screen "701_Line_Overview_1" 1280x800
   GraphicView "Graphic view_1" at 63,116 size 1157x650; Picture "b1 123927_1"
   Button "Template_Button_3" at 1074,2 size 203x55; TextOn 'FAULT RESET FAULT RESET'; TextOff 'FAULT RESET FAULT RESET'
      on Release: ResetBit("DB_SDC_GLOBAL_M.SDC_ER_Reset")
      on Press: SetBit("DB_SDC_GLOBAL_M.SDC_ER_Reset")
   AlarmView "Template_Alarm view_2" at 128,2 size 948x112
   Button "Template_Button_4" at 1196,56 size 81x59; TextOff 'Text'
      Appearance <- "AlwaysTRUE"
   Button "Button_7" at 0,57 size 128x58; TextOff 'SELECT SCREEN'
      on Release: ActivateScreen("010_START", 0)
   Button "Button_6" at 0,0 size 128x58; TextOff 'PREVIOUS SCREEN'
      on Click: function_efd93a16()
   DateTimeField "Template_Date/time field_2" at 1075,56 size 123x28
   DateTimeField "Template_Date/time field_3" at 1075,83 size 122x32
   TextField "Text field_1" at 981,345 size 46x25; Text 'S14'
   TextField "Text field_2" at 901,345 size 46x25; Text 'S13'
   TextField "Text field_3" at 818,344 size 46x25; Text 'S12'
   TextField "Text field_4" at 778,344 size 46x25; Text 'S11'
   TextField "Text field_5" at 734,344 size 46x25; Text 'S10'
   TextField "Text field_6" at 696,344 size 46x25; Text 'S9'
   TextField "Text field_7" at 653,344 size 46x25; Text 'S57'
   TextField "Text field_8" at 296,344 size 46x25; Text 'S7'
   TextField "Text field_9" at 252,344 size 46x25; Text 'S6'
   TextField "Text field_126" at 454,147 size 327x28; Text 'OVERVIEW 1 - SCREEN 701'
   TextField "Text field_130" at 23,313 size 82x24; Text 'EMS01R2'
   TextField "Text field_131" at 38,329 size 49x24; Text 'JB33'
   TextField "Text field_132" at 28,370 size 71x22; Text 'AREA A'
   TextField "Text field_10" at 135,418 size 46x25; Text 'S5'
   TextField "Text field_11" at 226,507 size 46x25; Text 'S4'
   TextField "Text field_12" at 133,473 size 46x25; Text 'S3'
   TextField "Text field_13" at 13,560 size 46x25; Text 'S2'
   TextField "Text field_14" at 4,640 size 46x25; Text 'S58'
   TextField "Text field_15" at 13,677 size 46x25; Text 'S1'
   TextField "Text field_16" at 5,716 size 46x25; Text 'S56'
   TextField "Text field_17" at 115,721 size 46x25; Text 'S55'
   TextField "Text field_18" at 116,560 size 71x22; Text 'AREA A'
   TextField "Text field_123" at 300,422 size 53x27; Text 'DL1'
   TextField "Text field_116" at 486,494 size 71x22; Text 'AREA G'
   TextField "Text field_119" at 508,426 size 82x22; Text 'AREA AA'
   TextField "Text field_127" at 607,453 size 82x24; Text 'EMS01R3'
   TextField "Text field_129" at 612,518 size 71x22; Text 'AREA B'
   TextField "Text field_19" at 606,485 size 82x22; Text 'AREA AA'
   TextField "Text field_121" at 731,425 size 53x27; Text 'DL2'
   TextField "Text field_122" at 712,450 size 93x25; Text 'Mrg Cell'
   TextField "Text field_120" at 948,425 size 71x22; Text 'AREA B'
   TextField "Text field_20" at 232,731 size 46x25; Text 'S54'
   TextField "Text field_21" at 195,612 size 46x25; Text 'S53'
   TextField "Text field_22" at 278,612 size 46x25; Text 'S52'
   TextField "Text field_23" at 348,613 size 46x25; Text 'S51'
   TextField "Text field_24" at 463,522 size 46x25; Text 'S47'
   TextField "Text field_25" at 534,521 size 46x25; Text 'S48'
   TextField "Text field_26" at 460,696 size 46x25; Text 'S44'
   TextField "Text field_27" at 529,696 size 46x25; Text 'S43'
   TextField "Text field_28" at 667,695 size 46x25; Text 'S42'
   TextField "Text field_29" at 719,657 size 46x25; Text 'S41'
   TextField "Text field_30" at 774,554 size 46x25; Text 'S40'
   TextField "Text field_31" at 883,638 size 46x25; Text 'S39'
   TextField "Text field_32" at 1015,638 size 46x25; Text 'S38'
   TextField "Text field_33" at 1114,638 size 46x25; Text 'S37'
   TextField "Text field_34" at 1158,533 size 46x25; Text 'S36'
   TextField "Text field_35" at 1157,469 size 46x25; Text 'S35'
   TextField "Text field_124" at 109,653 size 49x25; Text 'Cab'
   TextField "Text field_125" at 109,674 size 49x25; Text 'Pick'
   TextField "Text field_117" at 244,698 size 82x22; Text 'AREA FF'
   TextField "Text field_133" at 313,495 size 82x24; Text 'EMS01R1'
   TextField "Text field_134" at 319,518 size 71x22; Text 'AREA G'
   TextField "Text field_135" at 320,545 size 71x22; Text 'AREA F'
   TextField "Text field_136" at 314,570 size 82x22; Text 'AREA FF'
   TextField "Text field_137" at 785,680 size 60x24; Text 'EMS01'
   TextField "Text field_138" at 781,711 size 71x22; Text 'AREA D'
   TextField "Text field_139" at 781,739 size 71x22; Text 'AREA E'
   TextField "Text field_140" at 872,679 size 82x24; Text 'EMS01R4'
   TextField "Text field_143" at 979,672 size 60x24; Text 'EMS01'
   TextField "Text field_144" at 984,686 size 49x24; Text 'JB22'
   TextField "Text field_142" at 878,739 size 71x22; Text 'AREA H'
   TextField "Text field_146" at 973,738 size 71x22; Text 'AREA C'
   TextField "Text field_141" at 872,711 size 82x22; Text 'AREA CC'
   TextField "Text field_145" at 968,710 size 82x22; Text 'AREA BB'
   Button "Button_4" at 3,137 size 127x87; TextOn 'LINE_OVERVIEW_2 LINE OVERVIEW_2'; TextOff 'LINE_OVERVIEW_2 / Main Screen'
      on Click: ActivateScreen("010_START", 0)
   Button "Button_1" at 136,137 size 127x87; TextOn 'LINE_OVERVIEW_2 LINE OVERVIEW_2'; TextOff 'LINE_OVERVIEW_2 System Overview Screen'
      on Click: ActivateScreen("700_System_Line_Overview", 0)
   TextField "Text field_36" at 604,344 size 46x25; Text 'S8'
   Button "Button_2" at 0,0 size 37x32; TextOff 'Text'
      on Release: ActivateScreen("711_CARRIER_STATUS", 0)
      on Press: SetTag("HMI_EMS_Nr", "CarrierNumber")
   Button "Button_5" at 48,712 size 37x32; TextOff 'Text'
      on Release: ActivateScreen("711_CARRIER_STATUS", 0)
      on Press: SetTag("HMI_EMS_Nr", "CarrierNumber")
   Button "Button_8" at 116,760 size 37x32; TextOff 'Text'
      on Release: ActivateScreen("711_CARRIER_STATUS", 0)
      on Press: SetTag("HMI_EMS_Nr", "CarrierNumber")
   Button "Button_9" at 185,729 size 37x32; TextOff 'Text'
      on Release: ActivateScreen("711_CARRIER_STATUS", 0)
      on Press: SetTag("HMI_EMS_Nr", "CarrierNumber")
   Button "Button_10" at 186,691 size 37x32; TextOff 'Text'
      on Release: ActivateScreen("711_CARRIER_STATUS", 0)
      on Press: SetTag("HMI_EMS_Nr", "CarrierNumber")
   Button "Button_11" at 197,654 size 37x32; TextOff 'Text'
      on Release: ActivateScreen("711_CARRIER_STATUS", 0)
      on Press: SetTag("HMI_EMS_Nr", "CarrierNumber")
   Button "Button_12" at 238,654 size 37x32; TextOff 'Text'
      on Release: ActivateScreen("711_CARRIER_STATUS", 0)
      on Press: SetTag("HMI_EMS_Nr", "CarrierNumber")
   Button "Button_13" at 278,654 size 37x32; TextOff 'Text'
      on Release: ActivateScreen("711_CARRIER_STATUS", 0)
      on Press: SetTag("HMI_EMS_Nr", "CarrierNumber")
   Button "Button_14" at 316,654 size 37x32; TextOff 'Text'
      on Release: ActivateScreen("711_CARRIER_STATUS", 0)
      on Press: SetTag("HMI_EMS_Nr", "CarrierNumber")
   Button "Button_15" at 354,654 size 37x32; TextOff 'Text'
      on Release: ActivateScreen("711_CARRIER_STATUS", 0)
      on Press: SetTag("HMI_EMS_Nr", "CarrierNumber")
   Button "Button_16" at 461,654 size 37x32; TextOff 'Text'
      on Release: ActivateScreen("711_CARRIER_STATUS", 0)
      on Press: SetTag("HMI_EMS_Nr", "CarrierNumber")
   Button "Button_17" at 531,654 size 37x32; TextOff 'Text'
      on Release: ActivateScreen("711_CARRIER_STATUS", 0)
      on Press: SetTag("HMI_EMS_Nr", "CarrierNumber")
   Button "Button_18" at 630,654 size 37x32; TextOff 'Text'
      on Release: ActivateScreen("711_CARRIER_STATUS", 0)
      on Press: SetTag("HMI_EMS_Nr", "CarrierNumber")
   Button "Button_19" at 670,654 size 37x32; TextOff 'Text'
      on Release: ActivateScreen("711_CARRIER_STATUS", 0)
      on Press: SetTag("HMI_EMS_Nr", "CarrierNumber")
   Button "Button_20" at 723,623 size 37x32; TextOff 'Text'
      on Release: ActivateScreen("711_CARRIER_STATUS", 0)
      on Press: SetTag("HMI_EMS_Nr", "CarrierNumber")
   Button "Button_21" at 773,599 size 37x32; TextOff 'Text'
      on Release: ActivateScreen("711_CARRIER_STATUS", 0)
      on Press: SetTag("HMI_EMS_Nr", "CarrierNumber")
   Button "Button_22" at 813,599 size 37x32; TextOff 'Text'
      on Release: ActivateScreen("711_CARRIER_STATUS", 0)
      on Press: SetTag("HMI_EMS_Nr", "CarrierNumber")
   Button "Button_23" at 884,599 size 37x32; TextOff 'Text'
      on Release: ActivateScreen("711_CARRIER_STATUS", 0)
      on Press: SetTag("HMI_EMS_Nr", "CarrierNumber")
   Button "Button_24" at 924,599 size 37x32; TextOff 'Text'
      on Release: ActivateScreen("711_CARRIER_STATUS", 0)
      on Press: SetTag("HMI_EMS_Nr", "CarrierNumber")
   Button "Button_25" at 1014,599 size 37x32; TextOff 'Text'
      on Release: ActivateScreen("711_CARRIER_STATUS", 0)
      on Press: SetTag("HMI_EMS_Nr", "CarrierNumber")
   Button "Button_26" at 1054,599 size 37x32; TextOff 'Text'
      on Release: ActivateScreen("711_CARRIER_STATUS", 0)
      on Press: SetTag("HMI_EMS_Nr", "CarrierNumber")
   Button "Button_27" at 1115,599 size 37x32; TextOff 'Text'
      on Release: ActivateScreen("711_CARRIER_STATUS", 0)
      on Press: SetTag("HMI_EMS_Nr", "CarrierNumber")
   Button "Button_28" at 1156,599 size 37x32; TextOff 'Text'
      on Release: ActivateScreen("711_CARRIER_STATUS", 0)
      on Press: SetTag("HMI_EMS_Nr", "CarrierNumber")
   Button "Button_29" at 1218,529 size 37x32; TextOff 'Text'
      on Release: ActivateScreen("711_CARRIER_STATUS", 0)
      on Press: SetTag("HMI_EMS_Nr", "CarrierNumber")
   Button "Button_30" at 1219,466 size 37x32; TextOff 'Text'
      on Release: ActivateScreen("711_CARRIER_STATUS", 0)
      on Press: SetTag("HMI_EMS_Nr", "CarrierNumber")
   Button "Button_31" at 984,371 size 37x32; TextOff 'Text'
      on Release: ActivateScreen("711_CARRIER_STATUS", 0)
      on Press: SetTag("HMI_EMS_Nr", "CarrierNumber")
   Button "Button_32" at 945,371 size 37x32; TextOff 'Text'
      on Release: ActivateScreen("711_CARRIER_STATUS", 0)
      on Press: SetTag("HMI_EMS_Nr", "CarrierNumber")
   Button "Button_33" at 902,371 size 37x32; TextOff 'Text'
      on Release: ActivateScreen("711_CARRIER_STATUS", 0)
      on Press: SetTag("HMI_EMS_Nr", "CarrierNumber")
   Button "Button_34" at 863,371 size 37x32; TextOff 'Text'
      on Release: ActivateScreen("711_CARRIER_STATUS", 0)
      on Press: SetTag("HMI_EMS_Nr", "CarrierNumber")
   Button "Button_35" at 819,371 size 37x32; TextOff 'Text'
      on Release: ActivateScreen("711_CARRIER_STATUS", 0)
      on Press: SetTag("HMI_EMS_Nr", "CarrierNumber")
   Button "Button_36" at 778,371 size 37x32; TextOff 'Text'
      on Release: ActivateScreen("711_CARRIER_STATUS", 0)
      on Press: SetTag("HMI_EMS_Nr", "CarrierNumber")
   Button "Button_37" at 736,371 size 37x32; TextOff 'Text'
      on Release: ActivateScreen("711_CARRIER_STATUS", 0)
      on Press: SetTag("HMI_EMS_Nr", "CarrierNumber")
   Button "Button_38" at 692,371 size 37x32; TextOff 'Text'
      on Release: ActivateScreen("711_CARRIER_STATUS", 0)
      on Press: SetTag("HMI_EMS_Nr", "CarrierNumber")
   Button "Button_39" at 654,371 size 37x32; TextOff 'Text'
      on Release: ActivateScreen("711_CARRIER_STATUS", 0)
      on Press: SetTag("HMI_EMS_Nr", "CarrierNumber")
   Button "Button_40" at 610,371 size 37x32; TextOff 'Text'
      on Release: ActivateScreen("711_CARRIER_STATUS", 0)
      on Press: SetTag("HMI_EMS_Nr", "CarrierNumber")
   Button "Button_41" at 570,371 size 37x32; TextOff 'Text'
      on Release: ActivateScreen("711_CARRIER_STATUS", 0)
      on Press: SetTag("HMI_EMS_Nr", "CarrierNumber")
   Button "Button_42" at 530,371 size 37x32; TextOff 'Text'
      on Release: ActivateScreen("711_CARRIER_STATUS", 0)
      on Press: SetTag("HMI_EMS_Nr", "CarrierNumber")
   Button "Button_43" at 492,371 size 37x32; TextOff 'Text'
      on Release: ActivateScreen("711_CARRIER_STATUS", 0)
      on Press: SetTag("HMI_EMS_Nr", "CarrierNumber")
   Button "Button_44" at 453,371 size 37x32; TextOff 'Text'
      on Release: ActivateScreen("711_CARRIER_STATUS", 0)
      on Press: SetTag("HMI_EMS_Nr", "CarrierNumber")
   Button "Button_45" at 415,371 size 37x32; TextOff 'Text'
      on Release: ActivateScreen("711_CARRIER_STATUS", 0)
      on Press: SetTag("HMI_EMS_Nr", "CarrierNumber")
   Button "Button_46" at 376,371 size 37x32; TextOff 'Text'
      on Release: ActivateScreen("711_CARRIER_STATUS", 0)
      on Press: SetTag("HMI_EMS_Nr", "CarrierNumber")
   Button "Button_47" at 337,371 size 37x32; TextOff 'Text'
      on Release: ActivateScreen("711_CARRIER_STATUS", 0)
      on Press: SetTag("HMI_EMS_Nr", "CarrierNumber")
   Button "Button_48" at 292,371 size 37x32; TextOff 'Text'
      on Release: ActivateScreen("711_CARRIER_STATUS", 0)
      on Press: SetTag("HMI_EMS_Nr", "CarrierNumber")
   Button "Button_49" at 248,371 size 37x32; TextOff 'Text'
      on Release: ActivateScreen("711_CARRIER_STATUS", 0)
      on Press: SetTag("HMI_EMS_Nr", "CarrierNumber")
   Button "Button_50" at 172,414 size 37x32; TextOff 'Text'
      on Release: ActivateScreen("711_CARRIER_STATUS", 0)
      on Press: SetTag("HMI_EMS_Nr", "CarrierNumber")
   Button "Button_51" at 172,449 size 37x32; TextOff 'Text'
      on Release: ActivateScreen("711_CARRIER_STATUS", 0)
      on Press: SetTag("HMI_EMS_Nr", "CarrierNumber")
   Button "Button_52" at 171,503 size 37x32; TextOff 'Text'
      on Release: ActivateScreen("711_CARRIER_STATUS", 0)
      on Press: SetTag("HMI_EMS_Nr", "CarrierNumber")
   Button "Button_53" at 129,503 size 37x32; TextOff 'Text'
      on Release: ActivateScreen("711_CARRIER_STATUS", 0)
      on Press: SetTag("HMI_EMS_Nr", "CarrierNumber")
   TextField "Text field_37" at 579,695 size 46x25; Text 'S63'
   TextField "Text field_38" at 387,613 size 46x25; Text 'S45'
   Button "Button_59" at 584,654 size 37x32; TextOff 'Text'
      on Release: ActivateScreen("711_CARRIER_STATUS", 0)
      on Press: SetTag("HMI_EMS_Nr", "CarrierNumber")
   Group "Group" at 87,503 size 37x32
   Group "Group_1" at 47,596 size 37x32
   Group "Group_2" at 47,635 size 37x32
   Group "Group_3" at 47,672 size 37x32
   Group "Group_4" at 47,555 size 37x32; FormatPattern 99
   Button "Button_60" at 465,556 size 37x32; TextOff 'Text'
      on Release: ActivateScreen("711_CARRIER_STATUS", 0)
      on Press: SetTag("HMI_EMS_Nr", "CarrierNumber")
   Button "Button_61" at 535,556 size 37x32; TextOff 'Text'
      on Release: ActivateScreen("711_CARRIER_STATUS", 0)
      on Press: SetTag("HMI_EMS_Nr", "CarrierNumber")
   Button "Button_58" at 392,654 size 37x32; TextOff 'Text'
      on Release: ActivateScreen("711_CARRIER_STATUS", 0)
      on Press: SetTag("HMI_EMS_Nr", "CarrierNumber")
   IOField "I/O field_30" at 392,654 size 37x32; FormatPattern 99
      ProcessValue <- "CarrierNumber"
      Appearance <- "Faulted"
   IOField "I/O field_8" at 171,503 size 37x32; FormatPattern 99
      ProcessValue <- "CarrierNumber"
      Appearance <- "Faulted"
   IOField "I/O field_11" at 248,371 size 37x32; FormatPattern 99
      ProcessValue <- "CarrierNumber"
      Appearance <- "Faulted"
   IOField "I/O field_12" at 292,371 size 37x32; FormatPattern 99
      ProcessValue <- "CarrierNumber"
      Appearance <- "Faulted"
   IOField "I/O field_13" at 337,371 size 37x32; FormatPattern 99
      ProcessValue <- "CarrierNumber"
      Appearance <- "Faulted"
   IOField "I/O field_14" at 376,371 size 37x32; FormatPattern 99
      ProcessValue <- "CarrierNumber"
      Appearance <- "Faulted"
   IOField "I/O field_15" at 415,371 size 37x32; FormatPattern 99
      ProcessValue <- "CarrierNumber"
      Appearance <- "Faulted"
   IOField "I/O field_16" at 453,371 size 37x32; FormatPattern 99
      ProcessValue <- "CarrierNumber"
      Appearance <- "Faulted"
   IOField "I/O field_17" at 492,371 size 37x32; FormatPattern 99
      ProcessValue <- "CarrierNumber"
      Appearance <- "Faulted"
   IOField "I/O field_18" at 531,371 size 37x32; FormatPattern 99
      ProcessValue <- "CarrierNumber"
      Appearance <- "Faulted"
   IOField "I/O field_19" at 570,371 size 37x32; FormatPattern 99
      ProcessValue <- "CarrierNumber"
      Appearance <- "Faulted"
   IOField "I/O field_20" at 609,371 size 37x32; FormatPattern 99
      ProcessValue <- "CarrierNumber"
      Appearance <- "Faulted"
   IOField "I/O field_21" at 654,371 size 37x32; FormatPattern 99
      ProcessValue <- "CarrierNumber"
   IOField "I/O field_22" at 692,371 size 37x32; FormatPattern 99
      ProcessValue <- "CarrierNumber"
   IOField "I/O field_23" at 736,371 size 37x32; FormatPattern 99
      ProcessValue <- "CarrierNumber"
   IOField "I/O field_24" at 778,371 size 37x32; FormatPattern 99
      ProcessValue <- "CarrierNumber"
   IOField "I/O field_25" at 819,371 size 37x32; FormatPattern 99
      ProcessValue <- "CarrierNumber"
      Appearance <- "Faulted"
   IOField "I/O field_26" at 863,371 size 37x32; FormatPattern 99
      ProcessValue <- "CarrierNumber"
      Appearance <- "Faulted"
   IOField "I/O field_27" at 902,371 size 37x32; FormatPattern 99
      ProcessValue <- "CarrierNumber"
      Appearance <- "Faulted"
   IOField "I/O field_28" at 945,371 size 37x32; FormatPattern 99
      ProcessValue <- "CarrierNumber"
      Appearance <- "Faulted"
   IOField "I/O field_29" at 984,371 size 37x32; FormatPattern 99
      ProcessValue <- "CarrierNumber"
      Appearance <- "Faulted"
   IOField "I/O field_42" at 116,761 size 37x32; FormatPattern 99
      ProcessValue <- "CarrierNumber"
      Appearance <- "Faulted"
   IOField "I/O field_1" at 48,712 size 37x32; FormatPattern 99
      ProcessValue <- "CarrierNumber"
      Appearance <- "Faulted"
   IOField "I/O field_7" at 129,503 size 37x32; FormatPattern 99
      ProcessValue <- "CarrierNumber"
      Appearance <- "Faulted"
   IOField "I/O field_9" at 172,449 size 37x32; FormatPattern 99
      ProcessValue <- "CarrierNumber"
      Appearance <- "Faulted"
   IOField "I/O field_10" at 172,414 size 37x32; FormatPattern 99
      ProcessValue <- "CarrierNumber"
      Appearance <- "Faulted"
   IOField "I/O field_61" at 723,623 size 37x32; FormatPattern 99
      ProcessValue <- "CarrierNumber"
      Appearance <- "Faulted"
   IOField "I/O field_62" at 670,654 size 37x32; FormatPattern 99
      ProcessValue <- "CarrierNumber"
      Appearance <- "Faulted"
   IOField "I/O field_63" at 584,654 size 37x32; FormatPattern 99
      ProcessValue <- "CarrierNumber"
      Appearance <- "Faulted"
   IOField "I/O field_64" at 535,556 size 37x32; FormatPattern 99
      ProcessValue <- "CarrierNumber"
      Appearance <- "Faulted"
   IOField "I/O field_65" at 465,556 size 37x32; FormatPattern 99
      ProcessValue <- "CarrierNumber"
      Appearance <- "Faulted"
   IOField "I/O field_66" at 531,654 size 37x32; FormatPattern 99
      ProcessValue <- "CarrierNumber"
      Appearance <- "Faulted"
   IOField "I/O field_67" at 460,655 size 37x32; FormatPattern 99
      ProcessValue <- "CarrierNumber"
      Appearance <- "Faulted"
   IOField "I/O field_68" at 354,654 size 37x32; FormatPattern 99
      ProcessValue <- "CarrierNumber"
      Appearance <- "Faulted"
   IOField "I/O field_69" at 316,654 size 37x32; FormatPattern 99
      ProcessValue <- "CarrierNumber"
      Appearance <- "Faulted"
   IOField "I/O field_70" at 278,654 size 37x32; FormatPattern 99
      ProcessValue <- "CarrierNumber"
      Appearance <- "Faulted"
   IOField "I/O field_71" at 238,654 size 37x32; FormatPattern 99
      ProcessValue <- "CarrierNumber"
      Appearance <- "Faulted"
   IOField "I/O field_72" at 197,654 size 37x32; FormatPattern 99
      ProcessValue <- "CarrierNumber"
      Appearance <- "Faulted"
   IOField "I/O field_73" at 186,690 size 37x32; FormatPattern 99
      ProcessValue <- "CarrierNumber"
      Appearance <- "Faulted"
   IOField "I/O field_74" at 185,729 size 37x32; FormatPattern 99
      ProcessValue <- "CarrierNumber"
      Appearance <- "Faulted"
   IOField "I/O field_51" at 1219,466 size 37x32; FormatPattern 99
      ProcessValue <- "CarrierNumber"
      Appearance <- "Faulted"
   IOField "I/O field_52" at 1218,529 size 37x32; FormatPattern 99
      ProcessValue <- "CarrierNumber"
      Appearance <- "Faulted"
   IOField "I/O field_53" at 1156,599 size 37x32; FormatPattern 99
      ProcessValue <- "CarrierNumber"
      Appearance <- "Faulted"
   IOField "I/O field_54" at 1115,599 size 37x32; FormatPattern 99
      ProcessValue <- "CarrierNumber"
      Appearance <- "Faulted"
   IOField "I/O field_55" at 1054,599 size 37x32; FormatPattern 99
      ProcessValue <- "CarrierNumber"
      Appearance <- "Faulted"
   IOField "I/O field_56" at 1015,599 size 37x32; FormatPattern 99
      ProcessValue <- "CarrierNumber"
      Appearance <- "Faulted"
   IOField "I/O field_57" at 924,599 size 37x32; FormatPattern 99
      ProcessValue <- "CarrierNumber"
      Appearance <- "Faulted"
   IOField "I/O field_58" at 884,599 size 37x32; FormatPattern 99
      ProcessValue <- "CarrierNumber"
      Appearance <- "Faulted"
   IOField "I/O field_59" at 813,599 size 37x32; FormatPattern 99
      ProcessValue <- "CarrierNumber"
      Appearance <- "Faulted"
   IOField "I/O field_60" at 773,599 size 37x32; FormatPattern 99
      ProcessValue <- "CarrierNumber"
      Appearance <- "Faulted"
   IOField "I/O field_31" at 630,654 size 37x32; FormatPattern 99
      ProcessValue <- "CarrierNumber"
      Appearance <- "Faulted"
   Button "Button_54" at 87,503 size 37x32; TextOff 'Text'
      on Release: ActivateScreen("711_CARRIER_STATUS", 0)
      on Press: SetTag("HMI_EMS_Nr", "CarrierNumber")
   IOField "I/O field_6" at 87,503 size 37x32; FormatPattern 99
      ProcessValue <- "CarrierNumber"
      Appearance <- "Faulted"
   Button "Button_56" at 47,596 size 37x32; TextOff 'Text'
      on Release: ActivateScreen("711_CARRIER_STATUS", 0)
      on Press: SetTag("HMI_EMS_Nr", "CarrierNumber")
   IOField "I/O field_4" at 47,596 size 37x32; FormatPattern 99
      ProcessValue <- "CarrierNumber"
      Appearance <- "Faulted"
   Button "Button_57" at 47,635 size 37x32; TextOff 'Text'
      on Release: ActivateScreen("711_CARRIER_STATUS", 0)
      on Press: SetTag("HMI_EMS_Nr", "CarrierNumber")
   IOField "I/O field_3" at 47,635 size 37x32; FormatPattern 99
      ProcessValue <- "CarrierNumber"
      Appearance <- "Faulted"
   Button "Button_3" at 47,672 size 37x32; TextOff 'Text'
      on Release: ActivateScreen("711_CARRIER_STATUS", 0)
      on Press: SetTag("HMI_EMS_Nr", "CarrierNumber")
   IOField "I/O field_2" at 47,672 size 37x32; FormatPattern 99
      ProcessValue <- "CarrierNumber"
      Appearance <- "Faulted"
   Button "Button_55" at 47,555 size 37x32; TextOff 'Text'
      on Release: ActivateScreen("711_CARRIER_STATUS", 0)
      on Press: SetTag("HMI_EMS_Nr", "CarrierNumber")
   IOField "I/O field_5" at 47,555 size 37x32; FormatPattern 99999
      ProcessValue <- "CarrierNumber"
      Appearance <- "Faulted"

screen "702_Line_Overview_2" 1280x800
   Button "Template_Button_3" at 1074,2 size 203x55; TextOn 'FAULT RESET FAULT RESET'; TextOff 'FAULT RESET FAULT RESET'
      on Release: ResetBit("DB_SDC_GLOBAL_M.SDC_ER_Reset")
      on Press: SetBit("DB_SDC_GLOBAL_M.SDC_ER_Reset")
   AlarmView "Template_Alarm view_2" at 128,2 size 948x112
   Button "Template_Button_4" at 1196,56 size 81x59; TextOff 'Text'
      Appearance <- "AlwaysTRUE"
   Button "Button_7" at 0,57 size 128x58; TextOff 'SELECT SCREEN'
      on Release: ActivateScreen("010_START", 0)
   Button "Button_6" at 0,0 size 128x58; TextOff 'PREVIOUS SCREEN'
      on Click: function_efd93a16()
   DateTimeField "Template_Date/time field_2" at 1075,56 size 123x28
   DateTimeField "Template_Date/time field_3" at 1075,83 size 122x32
   TextField "Text field_2" at 485,123 size 341x28; Text 'OVERVIEW 2 - SCREEN 0024'
   GraphicView "Graphic view_1" at 250,117 size 646x682; Picture "Graphic_3"
   TextField "Text field_1" at 882,117 size 46x25; Text 'S16'
   TextField "Text field_3" at 882,152 size 46x25; Text 'S15'
   TextField "Text field_79" at 605,328 size 60x24; Text 'EMS01'
   TextField "Text field_80" at 608,342 size 49x24; Text 'JB22'
   TextField "Text field_81" at 592,369 size 82x22; Text 'AREA BB'
   TextField "Text field_4" at 477,123 size 327x28; Text 'OVERVIEW 2 - SCREEN 702'
   Button "Button_4" at 1148,702 size 127x87; TextOn 'LINE_OVERVIEW_2 LINE OVERVIEW_2'; TextOff 'LINE_OVERVIEW_2 / Main Screen'
      on Click: ActivateScreen("010_START", 0)
   Button "Button_1" at 1011,702 size 127x87; TextOn 'LINE_OVERVIEW_2 LINE OVERVIEW_2'; TextOff 'LINE_OVERVIEW_2 System Overview Screen'
      on Click: ActivateScreen("700_System_Line_Overview", 0)
   Button "Button_2" at 833,115 size 37x32; TextOff 'Text'
      on Release: ActivateScreen("711_CARRIER_STATUS", 0)
      on Press: SetTag("HMI_EMS_Nr", "CarrierNumber")
   Button "Button_3" at 833,147 size 37x32; TextOff 'Text'
      on Release: ActivateScreen("711_CARRIER_STATUS", 0)
      on Press: SetTag("HMI_EMS_Nr", "CarrierNumber")
   Button "Button_5" at 833,178 size 37x32; TextOff 'Text'
      on Release: ActivateScreen("711_CARRIER_STATUS", 0)
      on Press: SetTag("HMI_EMS_Nr", "CarrierNumber")
   Button "Button_8" at 833,209 size 37x32; TextOff 'Text'
      on Release: ActivateScreen("711_CARRIER_STATUS", 0)
      on Press: SetTag("HMI_EMS_Nr", "CarrierNumber")
   Button "Button_9" at 833,240 size 37x32; TextOff 'Text'
      on Release: ActivateScreen("711_CARRIER_STATUS", 0)
      on Press: SetTag("HMI_EMS_Nr", "CarrierNumber")
   Button "Button_10" at 833,273 size 37x32; TextOff 'Text'
      on Release: ActivateScreen("711_CARRIER_STATUS", 0)
      on Press: SetTag("HMI_EMS_Nr", "CarrierNumber")
   Button "Button_11" at 833,305 size 37x32; TextOff 'Text'
      on Release: ActivateScreen("711_CARRIER_STATUS", 0)
      on Press: SetTag("HMI_EMS_Nr", "CarrierNumber")
   Button "Button_12" at 833,337 size 37x32; TextOff 'Text'
      on Release: ActivateScreen("711_CARRIER_STATUS", 0)
      on Press: SetTag("HMI_EMS_Nr", "CarrierNumber")
   Button "Button_13" at 833,369 size 37x32; TextOff 'Text'
      on Release: ActivateScreen("711_CARRIER_STATUS", 0)
      on Press: SetTag("HMI_EMS_Nr", "CarrierNumber")
   Button "Button_14" at 833,401 size 37x32; TextOff 'Text'
      on Release: ActivateScreen("711_CARRIER_STATUS", 0)
      on Press: SetTag("HMI_EMS_Nr", "CarrierNumber")
   Button "Button_15" at 833,433 size 37x32; TextOff 'Text'
      on Release: ActivateScreen("711_CARRIER_STATUS", 0)
      on Press: SetTag("HMI_EMS_Nr", "CarrierNumber")
   Button "Button_16" at 833,464 size 37x32; TextOff 'Text'
      on Release: ActivateScreen("711_CARRIER_STATUS", 0)
      on Press: SetTag("HMI_EMS_Nr", "CarrierNumber")
   Button "Button_17" at 833,496 size 37x32; TextOff 'Text'
      on Release: ActivateScreen("711_CARRIER_STATUS", 0)
      on Press: SetTag("HMI_EMS_Nr", "CarrierNumber")
   Button "Button_18" at 833,528 size 37x32; TextOff 'Text'
      on Release: ActivateScreen("711_CARRIER_STATUS", 0)
      on Press: SetTag("HMI_EMS_Nr", "CarrierNumber")
   Button "Button_19" at 833,560 size 37x32; TextOff 'Text'
      on Release: ActivateScreen("711_CARRIER_STATUS", 0)
      on Press: SetTag("HMI_EMS_Nr", "CarrierNumber")
   Button "Button_20" at 833,592 size 37x32; TextOff 'Text'
      on Release: ActivateScreen("711_CARRIER_STATUS", 0)
      on Press: SetTag("HMI_EMS_Nr", "CarrierNumber")
   Button "Button_21" at 833,623 size 37x32; TextOff 'Text'
      on Release: ActivateScreen("711_CARRIER_STATUS", 0)
      on Press: SetTag("HMI_EMS_Nr", "CarrierNumber")
   Button "Button_22" at 833,654 size 37x32; TextOff 'Text'
      on Release: ActivateScreen("711_CARRIER_STATUS", 0)
      on Press: SetTag("HMI_EMS_Nr", "CarrierNumber")
   Button "Button_23" at 833,686 size 37x32; TextOff 'Text'
      on Release: ActivateScreen("711_CARRIER_STATUS", 0)
      on Press: SetTag("HMI_EMS_Nr", "CarrierNumber")
   Button "Button_24" at 833,718 size 37x32; TextOff 'Text'
      on Release: ActivateScreen("711_CARRIER_STATUS", 0)
      on Press: SetTag("HMI_EMS_Nr", "CarrierNumber")
   Button "Button_25" at 833,750 size 37x32; TextOff 'Text'
      on Release: ActivateScreen("711_CARRIER_STATUS", 0)
      on Press: SetTag("HMI_EMS_Nr", "CarrierNumber")
   IOField "I/O field_30" at 833,750 size 37x32; FormatPattern 99
      ProcessValue <- "CarrierNumber"
      Appearance <- "Faulted"
   IOField "I/O field_31" at 833,718 size 37x32; FormatPattern 99
      ProcessValue <- "CarrierNumber"
      Appearance <- "Faulted"
   IOField "I/O field_32" at 833,686 size 37x32; FormatPattern 99
      ProcessValue <- "CarrierNumber"
      Appearance <- "Faulted"
   IOField "I/O field_33" at 833,654 size 37x32; FormatPattern 99
      ProcessValue <- "CarrierNumber"
      Appearance <- "Faulted"
   IOField "I/O field_34" at 833,623 size 37x32; FormatPattern 99
      ProcessValue <- "CarrierNumber"
      Appearance <- "Faulted"
   IOField "I/O field_35" at 833,592 size 37x32; FormatPattern 99
      ProcessValue <- "CarrierNumber"
      Appearance <- "Faulted"
   IOField "I/O field_36" at 833,560 size 37x32; FormatPattern 99
      ProcessValue <- "CarrierNumber"
      Appearance <- "Faulted"
   IOField "I/O field_37" at 833,528 size 37x32; FormatPattern 99
      ProcessValue <- "CarrierNumber"
      Appearance <- "Faulted"
   IOField "I/O field_38" at 833,496 size 37x32; FormatPattern 99
      ProcessValue <- "CarrierNumber"
      Appearance <- "Faulted"
   IOField "I/O field_39" at 833,464 size 37x32; FormatPattern 99
      ProcessValue <- "CarrierNumber"
      Appearance <- "Faulted"
   IOField "I/O field_55" at 833,114 size 37x32; FormatPattern 99
      ProcessValue <- "CarrierNumber"
      Appearance <- "Faulted"
   IOField "I/O field_56" at 833,146 size 37x32; FormatPattern 99
      ProcessValue <- "CarrierNumber"
      Appearance <- "Faulted"
   IOField "I/O field_57" at 833,177 size 37x32; FormatPattern 99
      ProcessValue <- "CarrierNumber"
      Appearance <- "Faulted"
   IOField "I/O field_58" at 833,209 size 37x32; FormatPattern 99
      ProcessValue <- "CarrierNumber"
      Appearance <- "Faulted"
   IOField "I/O field_59" at 833,241 size 37x32; FormatPattern 99
      ProcessValue <- "CarrierNumber"
      Appearance <- "Faulted"
   IOField "I/O field_60" at 833,273 size 37x32; FormatPattern 99
      ProcessValue <- "CarrierNumber"
      Appearance <- "Faulted"
   IOField "I/O field_61" at 833,305 size 37x32; FormatPattern 99
      ProcessValue <- "CarrierNumber"
      Appearance <- "Faulted"
   IOField "I/O field_62" at 833,337 size 37x32; FormatPattern 99
      ProcessValue <- "CarrierNumber"
      Appearance <- "Faulted"
   IOField "I/O field_63" at 833,369 size 37x32; FormatPattern 99
      ProcessValue <- "CarrierNumber"
      Appearance <- "Faulted"
   IOField "I/O field_64" at 833,401 size 37x32; FormatPattern 99
      ProcessValue <- "CarrierNumber"
      Appearance <- "Faulted"
   IOField "I/O field_65" at 833,433 size 37x32; FormatPattern 99
      ProcessValue <- "CarrierNumber"
      Appearance <- "Faulted"

screen "703_Line_Overview_3" 1280x800
   Button "Template_Button_3" at 1074,2 size 203x55; TextOn 'FAULT RESET FAULT RESET'; TextOff 'FAULT RESET FAULT RESET'
      on Release: ResetBit("DB_SDC_GLOBAL_M.SDC_ER_Reset")
      on Press: SetBit("DB_SDC_GLOBAL_M.SDC_ER_Reset")
   AlarmView "Template_Alarm view_2" at 128,2 size 948x112
   Button "Template_Button_4" at 1196,56 size 81x59; TextOff 'Text'
      Appearance <- "AlwaysTRUE"
   Button "Button_7" at 0,57 size 128x58; TextOff 'SELECT SCREEN'
      on Release: ActivateScreen("010_START", 0)
   Button "Button_6" at 0,0 size 128x58; TextOff 'PREVIOUS SCREEN'
      on Click: function_efd93a16()
   DateTimeField "Template_Date/time field_2" at 1075,56 size 123x28
   DateTimeField "Template_Date/time field_3" at 1075,83 size 122x32
   GraphicView "Graphic view_1" at 26,247 size 1142x552; Picture "b2 124337_2"
   TextField "Text field_1" at 910,378 size 46x25; Text 'S17'
   TextField "Text field_15" at 77,290 size 46x25; Text 'S21'
   TextField "Text field_16" at 209,383 size 46x25; Text 'S20'
   TextField "Text field_17" at 612,381 size 46x25; Text 'S19'
   TextField "Text field_18" at 752,380 size 46x25; Text 'S18'
   TextField "Text field_5" at 1038,197 size 46x25; Text 'S32'
   TextField "Text field_6" at 828,197 size 46x25; Text 'S31'
   TextField "Text field_7" at 663,197 size 46x25; Text 'S30'
   TextField "Text field_8" at 577,197 size 46x25; Text 'S29'
   TextField "Text field_9" at 491,197 size 46x25; Text 'S28'
   TextField "Text field_10" at 414,197 size 46x25; Text 'S27'
   TextField "Text field_11" at 339,197 size 46x25; Text 'S26'
   TextField "Text field_12" at 277,163 size 46x25; Text 'S24'
   TextField "Text field_13" at 276,276 size 46x25; Text 'S23'
   TextField "Text field_14" at 211,198 size 46x25; Text 'S22'
   TextField "Text field_2" at 485,123 size 327x28; Text 'OVERVIEW 3 - SCREEN 703'
   TextField "Text field_4" at 1116,767 size 46x25; Text 'S33'
   TextField "Text field_79" at 1009,409 size 60x24; Text 'EMS01'
   TextField "Text field_80" at 1012,423 size 49x24; Text 'JB22'
   TextField "Text field_82" at 1002,461 size 71x22; Text 'AREA C'
   TextField "Text field_3" at 738,426 size 71x22; Text 'AREA C'
   TextField "Text field_76" at 379,430 size 82x24; Text 'EMS01R4'
   TextField "Text field_77" at 378,459 size 82x22; Text 'AREA CC'
   TextField "Text field_78" at 383,487 size 71x22; Text 'AREA H'
   TextField "Text field_73" at 123,291 size 82x22; Text 'AREA CC'
   TextField "Text field_121" at 489,285 size 61x28; Text 'DL5'
   TextField "Text field_72" at 926,291 size 71x22; Text 'AREA H'
   TextField "Text field_71" at 1077,550 size 71x22; Text 'AREA D'
   TextField "Text field_93" at 1008,626 size 60x24; Text 'EMS01'
   TextField "Text field_94" at 1003,660 size 71x22; Text 'AREA D'
   Button "Button_4" at 26,689 size 127x87; TextOn 'LINE_OVERVIEW_2 LINE OVERVIEW_2'; TextOff 'LINE_OVERVIEW_2 / Main Screen'
      on Click: ActivateScreen("010_START", 0)
   Button "Button_1" at 158,689 size 127x87; TextOn 'LINE_OVERVIEW_2 LINE OVERVIEW_2'; TextOff 'LINE_OVERVIEW_2 System Overview Screen'
      on Click: ActivateScreen("700_System_Line_Overview", 0)
   Button "Button_2" at 855,532 size 37x32; TextOff 'Text'
      on Release: ActivateScreen("711_CARRIER_STATUS", 0)
      on Press: SetTag("HMI_EMS_Nr", "CarrierNumber")
   Button "Button_3" at 855,500 size 37x32; TextOff 'Text'
      on Release: ActivateScreen("711_CARRIER_STATUS", 0)
      on Press: SetTag("HMI_EMS_Nr", "CarrierNumber")
   Button "Button_5" at 855,467 size 37x32; TextOff 'Text'
      on Release: ActivateScreen("711_CARRIER_STATUS", 0)
      on Press: SetTag("HMI_EMS_Nr", "CarrierNumber")
   Button "Button_8" at 855,435 size 37x32; TextOff 'Text'
      on Release: ActivateScreen("711_CARRIER_STATUS", 0)
      on Press: SetTag("HMI_EMS_Nr", "CarrierNumber")
   Button "Button_9" at 855,404 size 37x32; TextOff 'Text'
      on Release: ActivateScreen("711_CARRIER_STATUS", 0)
      on Press: SetTag("HMI_EMS_Nr", "CarrierNumber")
   Button "Button_10" at 855,372 size 37x32; TextOff 'Text'
      on Release: ActivateScreen("711_CARRIER_STATUS", 0)
      on Press: SetTag("HMI_EMS_Nr", "CarrierNumber")
   Button "Button_11" at 799,343 size 37x32; TextOff 'Text'
      on Release: ActivateScreen("711_CARRIER_STATUS", 0)
      on Press: SetTag("HMI_EMS_Nr", "CarrierNumber")
   Button "Button_12" at 753,343 size 37x32; TextOff 'Text'
      on Release: ActivateScreen("711_CARRIER_STATUS", 0)
      on Press: SetTag("HMI_EMS_Nr", "CarrierNumber")
   Button "Button_13" at 661,344 size 37x32; TextOff 'Text'
      on Release: ActivateScreen("711_CARRIER_STATUS", 0)
      on Press: SetTag("HMI_EMS_Nr", "CarrierNumber")
   Button "Button_14" at 613,344 size 37x32; TextOff 'Text'
      on Release: ActivateScreen("711_CARRIER_STATUS", 0)
      on Press: SetTag("HMI_EMS_Nr", "CarrierNumber")
   Button "Button_15" at 519,344 size 37x32; TextOff 'Text'
      on Release: ActivateScreen("711_CARRIER_STATUS", 0)
      on Press: SetTag("HMI_EMS_Nr", "CarrierNumber")
   Button "Button_16" at 475,344 size 37x32; TextOff 'Text'
      on Release: ActivateScreen("711_CARRIER_STATUS", 0)
      on Press: SetTag("HMI_EMS_Nr", "CarrierNumber")
   Button "Button_17" at 431,344 size 37x32; TextOff 'Text'
      on Release: ActivateScreen("711_CARRIER_STATUS", 0)
      on Press: SetTag("HMI_EMS_Nr", "CarrierNumber")
   Button "Button_18" at 387,344 size 37x32; TextOff 'Text'
      on Release: ActivateScreen("711_CARRIER_STATUS", 0)
      on Press: SetTag("HMI_EMS_Nr", "CarrierNumber")
   Button "Button_19" at 343,344 size 37x32; TextOff 'Text'
      on Release: ActivateScreen("711_CARRIER_STATUS", 0)
      on Press: SetTag("HMI_EMS_Nr", "CarrierNumber")
   Button "Button_20" at 299,344 size 37x32; TextOff 'Text'
      on Release: ActivateScreen("711_CARRIER_STATUS", 0)
      on Press: SetTag("HMI_EMS_Nr", "CarrierNumber")
   Button "Button_21" at 255,344 size 37x32; TextOff 'Text'
      on Release: ActivateScreen("711_CARRIER_STATUS", 0)
      on Press: SetTag("HMI_EMS_Nr", "CarrierNumber")
   Button "Button_22" at 211,344 size 37x32; TextOff 'Text'
      on Release: ActivateScreen("711_CARRIER_STATUS", 0)
      on Press: SetTag("HMI_EMS_Nr", "CarrierNumber")
   Button "Button_23" at 17,285 size 37x32; TextOff 'Text'
      on Release: ActivateScreen("711_CARRIER_STATUS", 0)
      on Press: SetTag("HMI_EMS_Nr", "CarrierNumber")
   Button "Button_24" at 122,230 size 37x32; TextOff 'Text'
      on Release: ActivateScreen("711_CARRIER_STATUS", 0)
      on Press: SetTag("HMI_EMS_Nr", "CarrierNumber")
   Button "Button_25" at 166,230 size 37x32; TextOff 'Text'
      on Release: ActivateScreen("711_CARRIER_STATUS", 0)
      on Press: SetTag("HMI_EMS_Nr", "CarrierNumber")
   Button "Button_26" at 212,230 size 37x32; TextOff 'Text'
      on Release: ActivateScreen("711_CARRIER_STATUS", 0)
      on Press: SetTag("HMI_EMS_Nr", "CarrierNumber")
   Button "Button_27" at 278,230 size 37x32; TextOff 'Text'
      on Release: ActivateScreen("711_CARRIER_STATUS", 0)
      on Press: SetTag("HMI_EMS_Nr", "CarrierNumber")
   Button "Button_28" at 342,230 size 37x32; TextOff 'Text'
      on Release: ActivateScreen("711_CARRIER_STATUS", 0)
      on Press: SetTag("HMI_EMS_Nr", "CarrierNumber")
   Button "Button_29" at 415,230 size 37x32; TextOff 'Text'
      on Release: ActivateScreen("711_CARRIER_STATUS", 0)
      on Press: SetTag("HMI_EMS_Nr", "CarrierNumber")
   Button "Button_30" at 279,193 size 37x32; TextOff 'Text'
      on Release: ActivateScreen("711_CARRIER_STATUS", 0)
      on Press: SetTag("HMI_EMS_Nr", "CarrierNumber")
   Button "Button_31" at 492,230 size 37x32; TextOff 'Text'
      on Release: ActivateScreen("711_CARRIER_STATUS", 0)
      on Press: SetTag("HMI_EMS_Nr", "CarrierNumber")
   Button "Button_32" at 578,230 size 37x32; TextOff 'Text'
      on Release: ActivateScreen("711_CARRIER_STATUS", 0)
      on Press: SetTag("HMI_EMS_Nr", "CarrierNumber")
   Button "Button_33" at 665,230 size 37x32; TextOff 'Text'
      on Release: ActivateScreen("711_CARRIER_STATUS", 0)
      on Press: SetTag("HMI_EMS_Nr", "CarrierNumber")
   Button "Button_34" at 768,230 size 37x32; TextOff 'Text'
      on Release: ActivateScreen("711_CARRIER_STATUS", 0)
      on Press: SetTag("HMI_EMS_Nr", "CarrierNumber")
   Button "Button_35" at 831,230 size 37x32; TextOff 'Text'
      on Release: ActivateScreen("711_CARRIER_STATUS", 0)
      on Press: SetTag("HMI_EMS_Nr", "CarrierNumber")
   Button "Button_36" at 974,230 size 37x32; TextOff 'Text'
      on Release: ActivateScreen("711_CARRIER_STATUS", 0)
      on Press: SetTag("HMI_EMS_Nr", "CarrierNumber")
   Button "Button_37" at 1041,230 size 37x32; TextOff 'Text'
      on Release: ActivateScreen("711_CARRIER_STATUS", 0)
      on Press: SetTag("HMI_EMS_Nr", "CarrierNumber")
   Button "Button_38" at 1174,267 size 37x32; TextOff 'Text'
      on Release: ActivateScreen("711_CARRIER_STATUS", 0)
      on Press: SetTag("HMI_EMS_Nr", "CarrierNumber")
   Button "Button_39" at 1174,300 size 37x32; TextOff 'Text'
      on Release: ActivateScreen("711_CARRIER_STATUS", 0)
      on Press: SetTag("HMI_EMS_Nr", "CarrierNumber")
   Button "Button_40" at 1174,333 size 37x32; TextOff 'Text'
      on Release: ActivateScreen("711_CARRIER_STATUS", 0)
      on Press: SetTag("HMI_EMS_Nr", "CarrierNumber")
   Button "Button_41" at 1174,366 size 37x32; TextOff 'Text'
      on Release: ActivateScreen("711_CARRIER_STATUS", 0)
      on Press: SetTag("HMI_EMS_Nr", "CarrierNumber")
   Button "Button_42" at 1174,399 size 37x32; TextOff 'Text'
      on Release: ActivateScreen("711_CARRIER_STATUS", 0)
      on Press: SetTag("HMI_EMS_Nr", "CarrierNumber")
   Button "Button_43" at 1174,432 size 37x32; TextOff 'Text'
      on Release: ActivateScreen("711_CARRIER_STATUS", 0)
      on Press: SetTag("HMI_EMS_Nr", "CarrierNumber")
   Button "Button_44" at 1174,465 size 37x32; TextOff 'Text'
      on Release: ActivateScreen("711_CARRIER_STATUS", 0)
      on Press: SetTag("HMI_EMS_Nr", "CarrierNumber")
   Button "Button_45" at 1174,498 size 37x32; TextOff 'Text'
      on Release: ActivateScreen("711_CARRIER_STATUS", 0)
      on Press: SetTag("HMI_EMS_Nr", "CarrierNumber")
   Button "Button_46" at 1174,531 size 37x32; TextOff 'Text'
      on Release: ActivateScreen("711_CARRIER_STATUS", 0)
      on Press: SetTag("HMI_EMS_Nr", "CarrierNumber")
   Button "Button_47" at 1174,564 size 37x32; TextOff 'Text'
      on Release: ActivateScreen("711_CARRIER_STATUS", 0)
      on Press: SetTag("HMI_EMS_Nr", "CarrierNumber")
   Button "Button_48" at 1174,597 size 37x32; TextOff 'Text'
      on Release: ActivateScreen("711_CARRIER_STATUS", 0)
      on Press: SetTag("HMI_EMS_Nr", "CarrierNumber")
   Button "Button_49" at 1174,630 size 37x32; TextOff 'Text'
      on Release: ActivateScreen("711_CARRIER_STATUS", 0)
      on Press: SetTag("HMI_EMS_Nr", "CarrierNumber")
   Button "Button_50" at 1174,663 size 37x32; TextOff 'Text'
      on Release: ActivateScreen("711_CARRIER_STATUS", 0)
      on Press: SetTag("HMI_EMS_Nr", "CarrierNumber")
   Button "Button_51" at 1174,696 size 37x32; TextOff 'Text'
      on Release: ActivateScreen("711_CARRIER_STATUS", 0)
      on Press: SetTag("HMI_EMS_Nr", "CarrierNumber")
   Button "Button_52" at 1174,729 size 37x32; TextOff 'Text'
      on Release: ActivateScreen("711_CARRIER_STATUS", 0)
      on Press: SetTag("HMI_EMS_Nr", "CarrierNumber")
   Button "Button_53" at 1174,762 size 37x32; TextOff 'Text'
      on Release: ActivateScreen("711_CARRIER_STATUS", 0)
      on Press: SetTag("HMI_EMS_Nr", "CarrierNumber")
   IOField "I/O field_3" at 17,285 size 37x32; FormatPattern 99
      ProcessValue <- "CarrierNumber"
      Appearance <- "Faulted"
   IOField "I/O field_37" at 211,344 size 37x32; FormatPattern 99
      ProcessValue <- "CarrierNumber"
      Appearance <- "Faulted"
   IOField "I/O field_38" at 255,344 size 37x32; FormatPattern 99
      ProcessValue <- "CarrierNumber"
      Appearance <- "Faulted"
   IOField "I/O field_39" at 299,344 size 37x32; FormatPattern 99
      ProcessValue <- "CarrierNumber"
      Appearance <- "Faulted"
   IOField "I/O field_40" at 343,344 size 37x32; FormatPattern 99
      ProcessValue <- "CarrierNumber"
      Appearance <- "Faulted"
   IOField "I/O field_41" at 387,344 size 37x32; FormatPattern 99
      ProcessValue <- "CarrierNumber"
      Appearance <- "Faulted"
   IOField "I/O field_42" at 431,344 size 37x32; FormatPattern 99
      ProcessValue <- "CarrierNumber"
      Appearance <- "Faulted"
   IOField "I/O field_43" at 475,344 size 37x32; FormatPattern 99
      ProcessValue <- "CarrierNumber"
      Appearance <- "Faulted"
   IOField "I/O field_44" at 519,344 size 37x32; FormatPattern 99
      ProcessValue <- "CarrierNumber"
      Appearance <- "Faulted"
   IOField "I/O field_45" at 613,344 size 37x32; FormatPattern 99
      ProcessValue <- "CarrierNumber"
      Appearance <- "Faulted"
   IOField "I/O field_46" at 661,344 size 37x32; FormatPattern 99
      ProcessValue <- "CarrierNumber"
      Appearance <- "Faulted"
   IOField "I/O field_47" at 753,343 size 37x32; FormatPattern 99
      ProcessValue <- "CarrierNumber"
      Appearance <- "Faulted"
   IOField "I/O field_48" at 799,343 size 37x32; FormatPattern 99
      ProcessValue <- "CarrierNumber"
      Appearance <- "Faulted"
   IOField "I/O field_49" at 855,372 size 37x32; FormatPattern 99
      ProcessValue <- "CarrierNumber"
      Appearance <- "Faulted"
   IOField "I/O field_50" at 855,404 size 37x32; FormatPattern 99
      ProcessValue <- "CarrierNumber"
      Appearance <- "Faulted"
   IOField "I/O field_51" at 855,436 size 37x32; FormatPattern 99
      ProcessValue <- "CarrierNumber"
      Appearance <- "Faulted"
   IOField "I/O field_52" at 855,468 size 37x32; FormatPattern 99
      ProcessValue <- "CarrierNumber"
      Appearance <- "Faulted"
   IOField "I/O field_53" at 855,500 size 37x32; FormatPattern 99
      ProcessValue <- "CarrierNumber"
      Appearance <- "Faulted"
   IOField "I/O field_54" at 855,532 size 37x32; FormatPattern 99
      ProcessValue <- "CarrierNumber"
      Appearance <- "Faulted"
   IOField "I/O field_1" at 279,230 size 37x32; FormatPattern 99
      ProcessValue <- "CarrierNumber"
      Appearance <- "Faulted"
   IOField "I/O field_2" at 166,230 size 37x32; FormatPattern 99
      ProcessValue <- "CarrierNumber"
      Appearance <- "Faulted"
   IOField "I/O field_4" at 212,230 size 37x32; FormatPattern 99
      ProcessValue <- "CarrierNumber"
      Appearance <- "Faulted"
   IOField "I/O field_5" at 279,193 size 37x32; FormatPattern 99
      ProcessValue <- "CarrierNumber"
      Appearance <- "Faulted"
   IOField "I/O field_6" at 122,230 size 37x32; FormatPattern 99
      ProcessValue <- "CarrierNumber"
      Appearance <- "Faulted"
   IOField "I/O field_7" at 342,230 size 37x32; FormatPattern 99
      ProcessValue <- "CarrierNumber"
      Appearance <- "Faulted"
   IOField "I/O field_8" at 415,230 size 37x32; FormatPattern 99
      ProcessValue <- "CarrierNumber"
      Appearance <- "Faulted"
   IOField "I/O field_9" at 492,230 size 37x32; FormatPattern 99
      ProcessValue <- "CarrierNumber"
      Appearance <- "Faulted"
   IOField "I/O field_10" at 578,230 size 37x32; FormatPattern 99
      ProcessValue <- "CarrierNumber"
      Appearance <- "Faulted"
   IOField "I/O field_11" at 665,230 size 37x32; FormatPattern 99
      ProcessValue <- "CarrierNumber"
      Appearance <- "Faulted"
   IOField "I/O field_12" at 768,230 size 37x32; FormatPattern 99
      ProcessValue <- "CarrierNumber"
      Appearance <- "Faulted"
   IOField "I/O field_13" at 831,230 size 37x32; FormatPattern 99
      ProcessValue <- "CarrierNumber"
      Appearance <- "Faulted"
   IOField "I/O field_14" at 974,230 size 37x32; FormatPattern 99
      ProcessValue <- "CarrierNumber"
      Appearance <- "Faulted"
   IOField "I/O field_15" at 1041,230 size 37x32; FormatPattern 99
      ProcessValue <- "CarrierNumber"
      Appearance <- "Faulted"
   IOField "I/O field_16" at 1174,267 size 37x32; FormatPattern 99
      ProcessValue <- "CarrierNumber"
      Appearance <- "Faulted"
   IOField "I/O field_17" at 1174,300 size 37x32; FormatPattern 99
      ProcessValue <- "CarrierNumber"
      Appearance <- "Faulted"
   IOField "I/O field_18" at 1174,333 size 37x32; FormatPattern 99
      ProcessValue <- "CarrierNumber"
      Appearance <- "Faulted"
   IOField "I/O field_19" at 1174,366 size 37x32; FormatPattern 99
      ProcessValue <- "CarrierNumber"
      Appearance <- "Faulted"
   IOField "I/O field_20" at 1174,399 size 37x32; FormatPattern 99
      ProcessValue <- "CarrierNumber"
      Appearance <- "Faulted"
   IOField "I/O field_21" at 1174,432 size 37x32; FormatPattern 99
      ProcessValue <- "CarrierNumber"
      Appearance <- "Faulted"
   IOField "I/O field_22" at 1174,465 size 37x32; FormatPattern 99
      ProcessValue <- "CarrierNumber"
      Appearance <- "Faulted"
   IOField "I/O field_23" at 1174,498 size 37x32; FormatPattern 99
      ProcessValue <- "CarrierNumber"
      Appearance <- "Faulted"
   IOField "I/O field_24" at 1174,531 size 37x32; FormatPattern 99
      ProcessValue <- "CarrierNumber"
      Appearance <- "Faulted"
   IOField "I/O field_25" at 1174,564 size 37x32; FormatPattern 99
      ProcessValue <- "CarrierNumber"
      Appearance <- "Faulted"
   IOField "I/O field_26" at 1174,597 size 37x32; FormatPattern 99
      ProcessValue <- "CarrierNumber"
      Appearance <- "Faulted"
   IOField "I/O field_27" at 1174,630 size 37x32; FormatPattern 99
      ProcessValue <- "CarrierNumber"
      Appearance <- "Faulted"
   IOField "I/O field_28" at 1174,663 size 37x32; FormatPattern 99
      ProcessValue <- "CarrierNumber"
      Appearance <- "Faulted"
   IOField "I/O field_29" at 1174,696 size 37x32; FormatPattern 99
      ProcessValue <- "CarrierNumber"
      Appearance <- "Faulted"
   IOField "I/O field_30" at 1174,729 size 37x32; FormatPattern 99
      ProcessValue <- "CarrierNumber"
      Appearance <- "Faulted"
   IOField "I/O field_31" at 1174,762 size 37x32; FormatPattern 99
      ProcessValue <- "CarrierNumber"
      Appearance <- "Faulted"